screen "St_Parameter" 320x240
   TextField "Text field_13" at 186,102 size 26x12; Text 'Hour'
   TextField "Text field_17" at 122,102 size 34x12; Text 'Second'
   TextField "Text field_10" at 118,88 size 86x16; Text 'Time Shift Setting'
   TextField "Text field_4" at 71,19 size 47x13; Text 'Day (1-31)'
   TextField "Text field_6" at 196,19 size 21x13; Text 'Year'
   TextField "Text field_5" at 119,19 size 61x12; Text 'Month (1-12)'
   TextField "Text field_1" at 6,1 size 143x17; Text 'STATISTIKA PARAMETER'
   TextField "Text field_2" at 9,32 size 62x15; Text 'Date Setting'
   TextField "Text field_3" at 10,65 size 61x15; Text 'Time Setting'
   TextField "Text field_7" at 67,54 size 52x12; Text 'Hour (0-23)'
   TextField "Text field_8" at 119,53 size 59x12; Text 'Minute (0-59)'
   TextField "Text field_9" at 176,53 size 64x12; Text 'Second (0-59)'
   IOField "I/O field_6" at 72,33 size 42x20; FormatPattern 99
      ProcessValue <- "DB_Integer_IDay"
   Button "Button_1" at 256,50 size 57x23; TextOff 'Execute'; TextOn 'OK'
      on Release: ResetBit("Data_Bool1_F_Set Time Day")
      on Press: SetBit("Data_Bool1_F_Set Time Day")
   TextField "Text field_11" at 11,117 size 33x15; Text 'Shift 1'
   TextField "Text field_15" at 49,102 size 26x12; Text 'Hour'
   TextField "Text field_16" at 85,102 size 30x12; Text 'Minute'
   IOField "I/O field_7" at 81,115 size 35x20; FormatPattern 99
      ProcessValue <- "DB_Integer_S1AMinute"
   IOField "I/O field_8" at 119,115 size 35x20; FormatPattern 99
      ProcessValue <- "DB_Integer_S1ASecond"
   TextField "Text field_12" at 160,114 size 17x15; Text 's/d'
   IOField "I/O field_9" at 180,115 size 35x20; FormatPattern 99
      ProcessValue <- "DB_Integer_S1BHour"
   TextField "Text field_14" at 221,102 size 30x12; Text 'Minute'
   TextField "Text field_18" at 256,102 size 34x12; Text 'Second'
   IOField "I/O field_11" at 218,115 size 35x20; FormatPattern 99
      ProcessValue <- "DB_Integer_S1BMinute"
   IOField "I/O field_12" at 256,115 size 35x20; FormatPattern 99
      ProcessValue <- "DB_Integer_S1BSecond"
   TextField "Text field_19" at 10,141 size 33x15; Text 'Shift 2'
   IOField "I/O field_13" at 43,139 size 35x20; FormatPattern 99
      ProcessValue <- "DB_Integer_S2AHour"
   IOField "I/O field_14" at 81,139 size 35x20; FormatPattern 99
      ProcessValue <- "DB_Integer_S2AMinute"
   IOField "I/O field_15" at 119,139 size 35x20; FormatPattern 99
      ProcessValue <- "DB_Integer_S2ASecond"
   TextField "Text field_23" at 160,140 size 17x15; Text 's/d'
   IOField "I/O field_16" at 180,139 size 35x20; FormatPattern 99
      ProcessValue <- "DB_Integer_S2BHour"
   IOField "I/O field_17" at 218,139 size 35x20; FormatPattern 99
      ProcessValue <- "DB_Integer_S2BMinute"
   IOField "I/O field_18" at 256,139 size 35x20; FormatPattern 99
      ProcessValue <- "DB_Integer_S2BSecond"
   TextField "Text field_27" at 9,165 size 33x15; Text 'Shift 3'
   IOField "I/O field_19" at 43,163 size 35x20; FormatPattern 99
      ProcessValue <- "DB_Integer_S3AHour"
   IOField "I/O field_20" at 81,163 size 35x20; FormatPattern 99
      ProcessValue <- "DB_Integer_S3AMinute"
   IOField "I/O field_21" at 119,163 size 35x20; FormatPattern 99
      ProcessValue <- "DB_Integer_S3ASecond"
   TextField "Text field_31" at 160,164 size 17x15; Text 's/d'
   IOField "I/O field_22" at 180,163 size 35x20; FormatPattern 99
      ProcessValue <- "DB_Integer_S3BHour"
   IOField "I/O field_23" at 218,163 size 35x20; FormatPattern 99
      ProcessValue <- "DB_Integer_S3BMinute"
   IOField "I/O field_24" at 256,163 size 35x20; FormatPattern 99
      ProcessValue <- "DB_Integer_S3BSecond"
   IOField "I/O field_10" at 43,115 size 35x20; FormatPattern 99
      ProcessValue <- "DB_Integer_S1AHour"
   IOField "I/O field_1" at 125,33 size 43x20; FormatPattern 99
      ProcessValue <- "DB_Integer_IMonth"
   IOField "I/O field_2" at 180,33 size 52x20; FormatPattern 9999
      ProcessValue <- "DB_Integer_IYear"
   IOField "I/O field_3" at 72,66 size 40x20; FormatPattern 99
      ProcessValue <- "DB_Integer_IHour"
   IOField "I/O field_4" at 129,66 size 40x20; FormatPattern 99
      ProcessValue <- "DB_Integer_IMinute"
   IOField "I/O field_5" at 185,66 size 40x20; FormatPattern 99
      ProcessValue <- "DB_Integer_ISecond"
   IOField "I/O field_25" at 163,1 size 155x23; FormatPattern 9999999999999999999999999999999999999999
      ProcessValue <- "Data_DTL1_Output"
   Button "Button_2" at 138,185 size 57x24; TextOff 'Execute'; TextOn 'OK'
   Button "Button_4" at 3,211 size 35x27; TextOff 'Main Page'; PictureOff "Home"
      on Click: ActivateScreen("Main Page", 0)

screen "Door Open Secret" 320x240
   Button "Button_1" at 100,205 size 120x30; TextOff 'Main Page'
      on Click: ActivateScreen("Main Page", 0)
   Switch "Switch_5" at 100,20 size 107x32; CaptionText 'Switch'; TextOff 'Safety Door On'; TextOn 'Safety Door Off'
      ProcessValue <- "Flag Enable/Disable Error Door Open"
   Switch "Switch_1" at 102,80 size 107x32; TextOff 'Reset'; CaptionText 'Switch'
      ProcessValue <- "AddReject2_DB_CountStop"
   IOField "I/O field_2" at 209,80 size 84x32; FormatPattern 999999999
      ProcessValue <- "AddReject2_DB_Countaddrej"

screen "St_Error Counter" 320x240
   TextField "Text field_13" at 244,51 size 70x129; Text 'Text'
   TextField "Text field_37" at 7,163 size 21x17; Text '8'
   IOField "I/O field_24" at 219,163 size 26x17; FormatPattern 999
      ProcessValue <- "Data_DTLData_DTL_Door Open[0].SECOND"
   IOField "I/O field_25" at 195,163 size 25x17; FormatPattern 999
      ProcessValue <- "Data_DTLData_DTL_Door Open[0].MINUTE"
   IOField "I/O field_26" at 171,163 size 25x17; FormatPattern 999
      ProcessValue <- "Data_DTLData_DTL_Door Open[0].HOUR"
   TextField "Text field_38" at 27,163 size 145x17; Text 'Door Open'
   IOField "I/O field_13" at 219,131 size 26x17; FormatPattern 999
      ProcessValue <- "Data_DTLData_DTL_Press Low[0].SECOND"
   IOField "I/O field_14" at 195,131 size 25x17; FormatPattern 999
      ProcessValue <- "Data_DTLData_DTL_Press Low[0].MINUTE"
   IOField "I/O field_15" at 171,131 size 25x17; FormatPattern 999
      ProcessValue <- "Data_DTLData_DTL_Press Low[0].HOUR"
   TextField "Text field_7" at 27,131 size 145x17; Text 'Pressure Low'
   TextField "Text field_35" at 7,147 size 21x17; Text '7'
   TextField "Text field_34" at 7,131 size 21x17; Text '6'
   TextField "Text field_33" at 7,115 size 21x17; Text '5'
   TextField "Text field_32" at 7,99 size 21x17; Text '4'
   TextField "Text field_31" at 7,83 size 21x17; Text '3'
   TextField "Text field_30" at 7,67 size 21x17; Text '2'
   TextField "Text field_29" at 7,51 size 21x17; Text '1'
   TextField "Text field_28" at 7,35 size 21x17; Text 'No'
   IOField "I/O field_8" at 219,147 size 26x17; FormatPattern 999
      ProcessValue <- "Data_DTLData_DTL_RS Pneu Er.SECOND"
   IOField "I/O field_16" at 195,147 size 25x17; FormatPattern 999
      ProcessValue <- "Data_DTLData_DTL_RS Pneu Er.MINUTE"
   IOField "I/O field_17" at 171,147 size 25x17; FormatPattern 999
      ProcessValue <- "Data_DTLData_DTL_RS Pneu Er.HOUR"
   IOField "I/O field_21" at 219,83 size 26x17; FormatPattern 999
      ProcessValue <- "Data_DTLData_DTL_Imaje Not In Position[0].SECOND"
   IOField "I/O field_22" at 195,83 size 25x17; FormatPattern 999
      ProcessValue <- "Data_DTLData_DTL_Imaje Not In Position[0].MINUTE"
   IOField "I/O field_23" at 171,83 size 25x17; FormatPattern 999
      ProcessValue <- "Data_DTLData_DTL_Imaje Not In Position[0].HOUR"
   TextField "Text field_25" at 27,83 size 145x17; Text 'Imaje Not In Position'
   IOField "I/O field_18" at 219,67 size 26x17; FormatPattern 999
      ProcessValue <- "Data_DTLData_DTL_Paper R Out[0].SECOND"
   IOField "I/O field_19" at 195,67 size 25x17; FormatPattern 999
      ProcessValue <- "Data_DTLData_DTL_Paper R Out[0].MINUTE"
   IOField "I/O field_20" at 171,67 size 25x17; FormatPattern 999
      ProcessValue <- "Data_DTLData_DTL_Paper R Out[0].HOUR"
   TextField "Text field_22" at 27,67 size 145x17; Text 'Imaje Paper Or Ribbon Out'
   TextField "Text field_2" at 171,35 size 25x17; Text 'Hour'
   IOField "I/O field_10" at 219,115 size 26x17; FormatPattern 999
      ProcessValue <- "Data_DTLData_DTL_Sloft Jam1.SECOND"
   IOField "I/O field_11" at 195,115 size 25x17; FormatPattern 999
      ProcessValue <- "Data_DTLData_DTL_Sloft Jam1.MINUTE"
   IOField "I/O field_12" at 171,115 size 25x17; FormatPattern 999
      ProcessValue <- "Data_DTLData_DTL_Sloft Jam1.HOUR"
   IOField "I/O field_4" at 219,99 size 26x17; FormatPattern 999
      ProcessValue <- "Data_DTLData_DTL_Always bad Read[0].SECOND"
   IOField "I/O field_5" at 195,99 size 25x17; FormatPattern 999
      ProcessValue <- "Data_DTLData_DTL_Always bad Read[0].MINUTE"
   IOField "I/O field_9" at 171,99 size 25x17; FormatPattern 999
      ProcessValue <- "Data_DTLData_DTL_Always bad Read[0].HOUR"
   TextField "Text field_12" at 219,35 size 26x17; Text 'Sec'
   TextField "Text field_11" at 195,35 size 25x17; Text 'Min'
   IOField "I/O field_2" at 219,51 size 26x17; FormatPattern 999
      ProcessValue <- "Data_DTLData_DTL_Imaje Er.SECOND"
   IOField "I/O field_1" at 195,51 size 25x17; FormatPattern 999
      ProcessValue <- "Data_DTLData_DTL_Imaje Er.MINUTE"
   TextField "Text field_3" at 27,35 size 145x17; Text 'Error Counter'
   TextField "Text field_4" at 27,51 size 145x17; Text 'System Imaje Error'
   TextField "Text field_5" at 27,99 size 145x17; Text 'Always Bad Read Sloft'
   IOField "I/O field_3" at 171,51 size 25x17; FormatPattern 999
      ProcessValue <- "Data_DTLData_DTL_Imaje Er.HOUR"
   TextField "Text field_9" at 120,17 size 18x13; Text 'S/D'
   TextField "Text field_1" at 3,0 size 197x18; Text 'CURRENT SHIFT (Error Counter)'
   TextField "Text field_36" at 260,0 size 57x15; Text 'Page 3 of 3'
   Button "Button_1" at 46,217 size 90x21; TextOff 'Statistic Data'
      on Click: ActivateScreen("St_Data Statistic", 0)
   Button "Button_3" at 1,218 size 41x20; TextOff 'Main Page'; PictureOff "Home"
      on Click: ActivateScreen("Main Page", 0)
   Button "Button_4" at 151,217 size 80x21; TextOff '<-- Back Page'; TextOn 'Page 2'
      on Click: ActivateScreen("St_Time machine data", 0)
   TextField "Text field_10" at 27,182 size 145x17; Text 'Downstream Jammed'
   IOField "I/O field_30" at 171,182 size 25x17; FormatPattern 999
      ProcessValue <- "Data_DTLData_DTL_Down Stop.HOUR"
   IOField "I/O field_31" at 195,182 size 25x17; FormatPattern 999
      ProcessValue <- "Data_DTLData_DTL_Down Stop.MINUTE"
   IOField "I/O field_32" at 219,182 size 26x17; FormatPattern 999
      ProcessValue <- "Data_DTLData_DTL_Down Stop.SECOND"
   TextField "Text field_14" at 244,182 size 70x17; Text 'Warning'
   IOField "I/O field_6" at 6,17 size 109x15; FormatPattern 9999999999999999999999999999999999999999
      ProcessValue <- "Data_DTL1_Cur_ShiftA"
   IOField "I/O field_7" at 143,17 size 109x15; FormatPattern 9999999999999999999999999999999999999999
      ProcessValue <- "Data_DTL1_Cur_ShiftB"
   TextField "Text field_15" at 263,115 size 7x15; Text ':'
   TextField "Text field_17" at 287,115 size 7x15; Text ':'
   IOField "I/O field_33" at 245,116 size 21x15; FormatPattern 999
      ProcessValue <- "Data_DTLData_DTL_Total Detail Error[0].HOUR"
   IOField "I/O field_34" at 268,116 size 21x15; FormatPattern 999
      ProcessValue <- "Data_DTLData_DTL_Total Detail Error[0].MINUTE"
   IOField "I/O field_35" at 291,116 size 21x15; FormatPattern 999
      ProcessValue <- "Data_DTLData_DTL_Total Detail Error[0].SECOND"
   TextField "Text field_16" at 244,35 size 70x17; Text 'Total (H:M:S)'
   TextField "Text field_8" at 27,115 size 145x17; Text 'Bundle Jammed'
   TextField "Text field_18" at 27,147 size 145x17; Text 'Reed Swicth pneumatic Error'
   IOField "I/O field_27" at 253,16 size 66x17; FormatPattern ????????
      ProcessValue <- "Data_String_sDT_Machine id"

screen "ST_Error Counter_1" 320x240
   TextField "Text field_13" at 244,51 size 70x129; Text 'Text'
   TextField "Text field_37" at 7,163 size 21x17; Text '8'
   IOField "I/O field_24" at 219,163 size 26x17; FormatPattern 999
      ProcessValue <- "Data_DTLData_DTL_Door Open[1].SECOND"
   IOField "I/O field_25" at 195,163 size 25x17; FormatPattern 999
      ProcessValue <- "Data_DTLData_DTL_Door Open[1].MINUTE"
   IOField "I/O field_26" at 171,163 size 25x17; FormatPattern 999
      ProcessValue <- "Data_DTLData_DTL_Door Open[1].HOUR"
   TextField "Text field_38" at 27,163 size 145x17; Text 'Door Open'
   IOField "I/O field_13" at 219,131 size 26x17; FormatPattern 999
      ProcessValue <- "Data_DTLData_DTL_Press Low[1].SECOND"
   IOField "I/O field_14" at 195,131 size 25x17; FormatPattern 999
      ProcessValue <- "Data_DTLData_DTL_Press Low[1].MINUTE"
   IOField "I/O field_15" at 171,131 size 25x17; FormatPattern 999
      ProcessValue <- "Data_DTLData_DTL_Press Low[1].HOUR"
   TextField "Text field_7" at 27,131 size 145x17; Text 'Pressure Low'
   TextField "Text field_35" at 7,147 size 21x17; Text '7'
   TextField "Text field_34" at 7,131 size 21x17; Text '6'
   TextField "Text field_33" at 7,115 size 21x17; Text '5'
   TextField "Text field_32" at 7,99 size 21x17; Text '4'
   TextField "Text field_31" at 7,83 size 21x17; Text '3'
   TextField "Text field_30" at 7,67 size 21x17; Text '2'
   TextField "Text field_29" at 7,51 size 21x17; Text '1'
   TextField "Text field_28" at 7,35 size 21x17; Text 'No'
   IOField "I/O field_8" at 219,147 size 26x17; FormatPattern 999
      ProcessValue <- "Data_DTLData_DTL_RS Pneu Er_1.SECOND"
   IOField "I/O field_16" at 195,147 size 25x17; FormatPattern 999
      ProcessValue <- "Data_DTLData_DTL_RS Pneu Er_1.MINUTE"
   IOField "I/O field_17" at 171,147 size 25x17; FormatPattern 999
      ProcessValue <- "Data_DTLData_DTL_RS Pneu Er_1.HOUR"
   IOField "I/O field_21" at 219,83 size 26x17; FormatPattern 999
      ProcessValue <- "Data_DTLData_DTL_Imaje Not In Position[1].SECOND"
   IOField "I/O field_22" at 195,83 size 25x17; FormatPattern 999
      ProcessValue <- "Data_DTLData_DTL_Imaje Not In Position[1].MINUTE"
   IOField "I/O field_23" at 171,83 size 25x17; FormatPattern 999
      ProcessValue <- "Data_DTLData_DTL_Imaje Not In Position[1].HOUR"
   TextField "Text field_25" at 27,83 size 145x17; Text 'Imaje Not In Position'
   IOField "I/O field_18" at 219,67 size 26x17; FormatPattern 999
      ProcessValue <- "Data_DTLData_DTL_Paper R Out[1].SECOND"
   IOField "I/O field_19" at 195,67 size 25x17; FormatPattern 999
      ProcessValue <- "Data_DTLData_DTL_Paper R Out[1].MINUTE"
   IOField "I/O field_20" at 171,67 size 25x17; FormatPattern 999
      ProcessValue <- "Data_DTLData_DTL_Paper R Out[1].HOUR"
   TextField "Text field_22" at 27,67 size 145x17; Text 'Imaje Paper Or Ribbon Out'
   TextField "Text field_2" at 171,35 size 25x17; Text 'Hour'
   IOField "I/O field_10" at 219,115 size 26x17; FormatPattern 999
      ProcessValue <- "Data_DTLData_DTL_Sloft Jam1_1.SECOND"
   IOField "I/O field_11" at 195,115 size 25x17; FormatPattern 999
      ProcessValue <- "Data_DTLData_DTL_Sloft Jam1_1.MINUTE"
   IOField "I/O field_12" at 171,115 size 25x17; FormatPattern 999
      ProcessValue <- "Data_DTLData_DTL_Sloft Jam1_1.HOUR"
   IOField "I/O field_4" at 219,99 size 26x17; FormatPattern 999
      ProcessValue <- "Data_DTLData_DTL_Always bad Read[1].SECOND"
   IOField "I/O field_5" at 195,99 size 25x17; FormatPattern 999
      ProcessValue <- "Data_DTLData_DTL_Always bad Read[1].MINUTE"
   IOField "I/O field_9" at 171,99 size 25x17; FormatPattern 999
      ProcessValue <- "Data_DTLData_DTL_Always bad Read[1].HOUR"
   TextField "Text field_12" at 219,35 size 26x17; Text 'Sec'
   TextField "Text field_11" at 195,35 size 25x17; Text 'Min'
   IOField "I/O field_2" at 219,51 size 26x17; FormatPattern 999
      ProcessValue <- "Data_DTLData_DTL_Imaje Er_1.SECOND"
   IOField "I/O field_1" at 195,51 size 25x17; FormatPattern 999
      ProcessValue <- "Data_DTLData_DTL_Imaje Er_1.MINUTE"
   TextField "Text field_3" at 27,35 size 145x17; Text 'Error Counter'
   TextField "Text field_4" at 27,51 size 145x17; Text 'System Imaje Error'
   TextField "Text field_5" at 27,99 size 145x17; Text 'Always Bad Read Sloft'
   IOField "I/O field_3" at 171,51 size 25x17; FormatPattern 999
      ProcessValue <- "Data_DTLData_DTL_Imaje Er_1.HOUR"
   TextField "Text field_9" at 120,17 size 18x13; Text 'S/D'
   TextField "Text field_1" at 3,0 size 159x18; Text 'CURRENT SHIFT MINUS 1'
   TextField "Text field_36" at 260,0 size 57x15; Text 'Page 3 of 3'
   Button "Button_1" at 46,217 size 90x21; TextOff 'Statistic Data'
      on Click: ActivateScreen("St_Data Statistic", 0)
   Button "Button_3" at 1,218 size 41x20; TextOff 'Main Page'; PictureOff "Home"
      on Click: ActivateScreen("Main Page", 0)
   Button "Button_4" at 151,217 size 80x21; TextOff '<-- Back Page'; TextOn 'Page 2'
      on Click: ActivateScreen("St_Time machine data_1", 0)
   TextField "Text field_10" at 27,182 size 145x17; Text 'Downstream Jammed'
   IOField "I/O field_30" at 171,182 size 25x17; FormatPattern 999
      ProcessValue <- "Data_DTLData_DTL_Down Stop_1.HOUR"
   IOField "I/O field_31" at 195,182 size 25x17; FormatPattern 999
      ProcessValue <- "Data_DTLData_DTL_Down Stop_1.MINUTE"
   IOField "I/O field_32" at 219,182 size 26x17; FormatPattern 999
      ProcessValue <- "Data_DTLData_DTL_Down Stop_1.SECOND"
   TextField "Text field_14" at 244,182 size 70x17; Text 'Warning'
   IOField "I/O field_7" at 143,17 size 109x15; FormatPattern 9999999999999999999999999999999999999999
      ProcessValue <- "Data_DTL1_Cur_ShiftB_1"
   IOField "I/O field_6" at 6,17 size 109x15; FormatPattern 9999999999999999999999999999999999999999
      ProcessValue <- "Data_DTL1_Cur_ShiftA_1"
   TextField "Text field_15" at 263,115 size 7x15; Text ':'
   TextField "Text field_17" at 287,115 size 7x15; Text ':'
   IOField "I/O field_33" at 245,116 size 21x15; FormatPattern 999
      ProcessValue <- "Data_DTLData_DTL_Total Detail Error[1].HOUR"
   IOField "I/O field_34" at 268,116 size 21x15; FormatPattern 999
      ProcessValue <- "Data_DTLData_DTL_Total Detail Error[1].MINUTE"
   IOField "I/O field_35" at 291,116 size 21x15; FormatPattern 999
      ProcessValue <- "Data_DTLData_DTL_Total Detail Error[1].SECOND"
   TextField "Text field_16" at 244,35 size 70x17; Text 'Total (H:M:S)'
   TextField "Text field_8" at 27,115 size 145x17; Text 'Bundle Jammed'
   TextField "Text field_18" at 27,147 size 145x17; Text 'Reed Swicth pneumatic Error'
   IOField "I/O field_27" at 253,16 size 66x17; FormatPattern ????????
      ProcessValue <- "Data_String_sDT_Machine id"

screen "St_Error Counter_2" 320x240
   TextField "Text field_13" at 244,51 size 70x129; Text 'Text'
   TextField "Text field_37" at 7,163 size 21x17; Text '8'
   IOField "I/O field_24" at 219,163 size 26x17; FormatPattern 999
      ProcessValue <- "Data_DTLData_DTL_Door Open[2].SECOND"
   IOField "I/O field_25" at 195,163 size 25x17; FormatPattern 999
      ProcessValue <- "Data_DTLData_DTL_Door Open[2].MINUTE"
   IOField "I/O field_26" at 171,163 size 25x17; FormatPattern 999
      ProcessValue <- "Data_DTLData_DTL_Door Open[2].HOUR"
   TextField "Text field_38" at 27,163 size 145x17; Text 'Door Open'
   IOField "I/O field_13" at 219,131 size 26x17; FormatPattern 999
      ProcessValue <- "Data_DTLData_DTL_Press Low[2].SECOND"
   IOField "I/O field_14" at 195,131 size 25x17; FormatPattern 999
      ProcessValue <- "Data_DTLData_DTL_Press Low[2].MINUTE"
   IOField "I/O field_15" at 171,131 size 25x17; FormatPattern 999
      ProcessValue <- "Data_DTLData_DTL_Press Low[2].HOUR"
   TextField "Text field_7" at 27,131 size 145x17; Text 'Pressure Low'
   TextField "Text field_35" at 7,147 size 21x17; Text '7'
   TextField "Text field_34" at 7,131 size 21x17; Text '6'
   TextField "Text field_33" at 7,115 size 21x17; Text '5'
   TextField "Text field_32" at 7,99 size 21x17; Text '4'
   TextField "Text field_31" at 7,83 size 21x17; Text '3'
   TextField "Text field_30" at 7,67 size 21x17; Text '2'
   TextField "Text field_29" at 7,51 size 21x17; Text '1'
   TextField "Text field_28" at 7,35 size 21x17; Text 'No'
   IOField "I/O field_8" at 219,147 size 26x17; FormatPattern 999
      ProcessValue <- "Data_DTLData_DTL_RS Pneu Er_2.SECOND"
   IOField "I/O field_16" at 195,147 size 25x17; FormatPattern 999
      ProcessValue <- "Data_DTLData_DTL_RS Pneu Er_2.MINUTE"
   IOField "I/O field_17" at 171,147 size 25x17; FormatPattern 999
      ProcessValue <- "Data_DTLData_DTL_RS Pneu Er_2.HOUR"
   IOField "I/O field_21" at 219,83 size 26x17; FormatPattern 999
      ProcessValue <- "Data_DTLData_DTL_Imaje Not In Position[2].SECOND"
   IOField "I/O field_22" at 195,83 size 25x17; FormatPattern 999
      ProcessValue <- "Data_DTLData_DTL_Imaje Not In Position[2].MINUTE"
   IOField "I/O field_23" at 171,83 size 25x17; FormatPattern 999
      ProcessValue <- "Data_DTLData_DTL_Imaje Not In Position[2].HOUR"
   TextField "Text field_25" at 27,83 size 145x17; Text 'Imaje Not In Position'
   IOField "I/O field_18" at 219,67 size 26x17; FormatPattern 999
      ProcessValue <- "Data_DTLData_DTL_Paper R Out[2].SECOND"
   IOField "I/O field_19" at 195,67 size 25x17; FormatPattern 999
      ProcessValue <- "Data_DTLData_DTL_Paper R Out[2].MINUTE"
   IOField "I/O field_20" at 171,67 size 25x17; FormatPattern 999
      ProcessValue <- "Data_DTLData_DTL_Paper R Out[2].HOUR"
   TextField "Text field_22" at 27,67 size 145x17; Text 'Imaje Paper Or Ribbon Out'
   TextField "Text field_2" at 171,35 size 25x17; Text 'Hour'
   IOField "I/O field_10" at 219,115 size 26x17; FormatPattern 999
      ProcessValue <- "Data_DTLData_DTL_Sloft Jam1_2.SECOND"
   IOField "I/O field_11" at 195,115 size 25x17; FormatPattern 999
      ProcessValue <- "Data_DTLData_DTL_Sloft Jam1_2.MINUTE"
   IOField "I/O field_12" at 171,115 size 25x17; FormatPattern 999
      ProcessValue <- "Data_DTLData_DTL_Sloft Jam1_2.HOUR"
   IOField "I/O field_4" at 219,99 size 26x17; FormatPattern 999
      ProcessValue <- "Data_DTLData_DTL_Always bad Read[2].SECOND"
   IOField "I/O field_5" at 195,99 size 25x17; FormatPattern 999
      ProcessValue <- "Data_DTLData_DTL_Always bad Read[2].MINUTE"
   IOField "I/O field_9" at 171,99 size 25x17; FormatPattern 999
      ProcessValue <- "Data_DTLData_DTL_Always bad Read[2].HOUR"
   TextField "Text field_12" at 219,35 size 26x17; Text 'Sec'
   TextField "Text field_11" at 195,35 size 25x17; Text 'Min'
   IOField "I/O field_2" at 219,51 size 26x17; FormatPattern 999
      ProcessValue <- "Data_DTLData_DTL_Imaje Er_2.SECOND"
   IOField "I/O field_1" at 195,51 size 25x17; FormatPattern 999
      ProcessValue <- "Data_DTLData_DTL_Imaje Er_2.MINUTE"
   TextField "Text field_3" at 27,35 size 145x17; Text 'Error Counter'
   TextField "Text field_4" at 27,51 size 145x17; Text 'System Imaje Error'
   TextField "Text field_5" at 27,99 size 145x17; Text 'Always Bad Read Sloft'
   IOField "I/O field_3" at 171,51 size 25x17; FormatPattern 999
      ProcessValue <- "Data_DTLData_DTL_Imaje Er_2.HOUR"
   IOField "I/O field_6" at 6,17 size 109x15; FormatPattern 9999999999999999999999999999999999999999
      ProcessValue <- "Data_DTL1_Cur_ShiftA_2"
   TextField "Text field_9" at 120,17 size 18x13; Text 'S/D'
   IOField "I/O field_7" at 143,17 size 109x15; FormatPattern 9999999999999999999999999999999999999999
      ProcessValue <- "Data_DTL1_Cur_ShiftB_2"
   TextField "Text field_1" at 3,0 size 159x18; Text 'CURRENT SHIFT MINUS 2'
   TextField "Text field_36" at 260,0 size 57x15; Text 'Page 3 of 3'
   Button "Button_1" at 46,217 size 90x21; TextOff 'Statistic Data'
      on Click: ActivateScreen("St_Data Statistic", 0)
   Button "Button_3" at 1,218 size 41x20; TextOff 'Main Page'; PictureOff "Home"
      on Click: ActivateScreen("Main Page", 0)
   Button "Button_4" at 151,217 size 80x21; TextOff '<-- Back Page'; TextOn 'Page 2'
      on Click: ActivateScreen("St_Time machine data_2", 0)
   TextField "Text field_10" at 27,182 size 145x17; Text 'Downstream Jammed'
   IOField "I/O field_30" at 171,182 size 25x17; FormatPattern 999
      ProcessValue <- "Data_DTLData_DTL_Down Stop_2.HOUR"
   IOField "I/O field_31" at 195,182 size 25x17; FormatPattern 999
      ProcessValue <- "Data_DTLData_DTL_Down Stop_2.MINUTE"
   IOField "I/O field_32" at 219,182 size 26x17; FormatPattern 999
      ProcessValue <- "Data_DTLData_DTL_Down Stop_2.SECOND"
   TextField "Text field_14" at 244,182 size 70x17; Text 'Warning'
   TextField "Text field_15" at 263,115 size 7x15; Text ':'
   TextField "Text field_17" at 287,115 size 7x15; Text ':'
   IOField "I/O field_33" at 245,116 size 21x15; FormatPattern 999
      ProcessValue <- "Data_DTLData_DTL_Total Detail Error[2].HOUR"
   IOField "I/O field_34" at 268,116 size 21x15; FormatPattern 999
      ProcessValue <- "Data_DTLData_DTL_Total Detail Error[2].MINUTE"
   IOField "I/O field_35" at 291,116 size 21x15; FormatPattern 999
      ProcessValue <- "Data_DTLData_DTL_Total Detail Error[2].SECOND"
   TextField "Text field_16" at 244,35 size 70x17; Text 'Total (H:M:S)'
   TextField "Text field_8" at 27,115 size 145x17; Text 'Bundle Jammed'
   TextField "Text field_18" at 27,147 size 145x17; Text 'Reed Swicth pneumatic Error'
   IOField "I/O field_27" at 253,16 size 66x17; FormatPattern ????????
      ProcessValue <- "Data_String_sDT_Machine id"

screen "St_Error Counter_3" 320x240
   TextField "Text field_13" at 244,51 size 70x129; Text 'Text'
   TextField "Text field_37" at 7,163 size 21x17; Text '8'
   IOField "I/O field_24" at 219,163 size 26x17; FormatPattern 999
      ProcessValue <- "Data_DTLData_DTL_Door Open[3].SECOND"
   IOField "I/O field_25" at 195,163 size 25x17; FormatPattern 999
      ProcessValue <- "Data_DTLData_DTL_Door Open[3].MINUTE"
   IOField "I/O field_26" at 171,163 size 25x17; FormatPattern 999
      ProcessValue <- "Data_DTLData_DTL_Door Open[3].HOUR"
   TextField "Text field_38" at 27,163 size 145x17; Text 'Door Open'
   IOField "I/O field_13" at 219,131 size 26x17; FormatPattern 999
      ProcessValue <- "Data_DTLData_DTL_Press Low[3].SECOND"
   IOField "I/O field_14" at 195,131 size 25x17; FormatPattern 999
      ProcessValue <- "Data_DTLData_DTL_Press Low[3].MINUTE"
   IOField "I/O field_15" at 171,131 size 25x17; FormatPattern 999
      ProcessValue <- "Data_DTLData_DTL_Press Low[3].HOUR"
   TextField "Text field_7" at 27,131 size 145x17; Text 'Pressure Low'
   TextField "Text field_35" at 7,147 size 21x17; Text '7'
   TextField "Text field_34" at 7,131 size 21x17; Text '6'
   TextField "Text field_33" at 7,115 size 21x17; Text '5'
   TextField "Text field_32" at 7,99 size 21x17; Text '4'
   TextField "Text field_31" at 7,83 size 21x17; Text '3'
   TextField "Text field_30" at 7,67 size 21x17; Text '2'
   TextField "Text field_29" at 7,51 size 21x17; Text '1'
   TextField "Text field_28" at 7,35 size 21x17; Text 'No'
   IOField "I/O field_8" at 219,147 size 26x17; FormatPattern 999
      ProcessValue <- "Data_DTLData_DTL_RS Pneu Er_3.SECOND"
   IOField "I/O field_16" at 195,147 size 25x17; FormatPattern 999
      ProcessValue <- "Data_DTLData_DTL_RS Pneu Er_3.MINUTE"
   IOField "I/O field_17" at 171,147 size 25x17; FormatPattern 999
      ProcessValue <- "Data_DTLData_DTL_RS Pneu Er_3.HOUR"
   IOField "I/O field_21" at 219,83 size 26x17; FormatPattern 999
      ProcessValue <- "Data_DTLData_DTL_Imaje Not In Position[3].SECOND"
   IOField "I/O field_22" at 195,83 size 25x17; FormatPattern 999
      ProcessValue <- "Data_DTLData_DTL_Imaje Not In Position[3].MINUTE"
   IOField "I/O field_23" at 171,83 size 25x17; FormatPattern 999
      ProcessValue <- "Data_DTLData_DTL_Imaje Not In Position[3].HOUR"
   TextField "Text field_25" at 27,83 size 145x17; Text 'Imaje Not In Position'
   IOField "I/O field_18" at 219,67 size 26x17; FormatPattern 999
      ProcessValue <- "Data_DTLData_DTL_Paper R Out[3].SECOND"
   IOField "I/O field_19" at 195,67 size 25x17; FormatPattern 999
      ProcessValue <- "Data_DTLData_DTL_Paper R Out[3].MINUTE"
   IOField "I/O field_20" at 171,67 size 25x17; FormatPattern 999
      ProcessValue <- "Data_DTLData_DTL_Paper R Out[3].HOUR"
   TextField "Text field_22" at 27,67 size 145x17; Text 'Imaje Paper Or Ribbon Out'
   TextField "Text field_2" at 171,35 size 25x17; Text 'Hour'
   IOField "I/O field_10" at 219,115 size 26x17; FormatPattern 999
      ProcessValue <- "Data_DTLData_DTL_Sloft Jam1_3.SECOND"
   IOField "I/O field_11" at 195,115 size 25x17; FormatPattern 999
      ProcessValue <- "Data_DTLData_DTL_Sloft Jam1_3.MINUTE"
   IOField "I/O field_12" at 171,115 size 25x17; FormatPattern 999
      ProcessValue <- "Data_DTLData_DTL_Sloft Jam1_3.HOUR"
   IOField "I/O field_4" at 219,99 size 26x17; FormatPattern 999
      ProcessValue <- "Data_DTLData_DTL_Always bad Read[3].SECOND"
   IOField "I/O field_5" at 195,99 size 25x17; FormatPattern 999
      ProcessValue <- "Data_DTLData_DTL_Always bad Read[3].MINUTE"
   IOField "I/O field_9" at 171,99 size 25x17; FormatPattern 999
      ProcessValue <- "Data_DTLData_DTL_Always bad Read[3].HOUR"
   TextField "Text field_12" at 219,35 size 26x17; Text 'Sec'
   TextField "Text field_11" at 195,35 size 25x17; Text 'Min'
   IOField "I/O field_2" at 219,51 size 26x17; FormatPattern 999
      ProcessValue <- "Data_DTLData_DTL_Imaje Er_3.SECOND"
   IOField "I/O field_1" at 195,51 size 25x17; FormatPattern 999
      ProcessValue <- "Data_DTLData_DTL_Imaje Er_3.MINUTE"
   TextField "Text field_3" at 27,35 size 145x17; Text 'Error Counter'
   TextField "Text field_4" at 27,51 size 145x17; Text 'System Imaje Error'
   TextField "Text field_5" at 27,99 size 145x17; Text 'Always Bad Read Sloft'
   IOField "I/O field_3" at 171,51 size 25x17; FormatPattern 999
      ProcessValue <- "Data_DTLData_DTL_Imaje Er_3.HOUR"
   IOField "I/O field_6" at 6,17 size 109x15; FormatPattern 9999999999999999999999999999999999999999
      ProcessValue <- "Data_DTL1_Cur_ShiftA_3"
   TextField "Text field_9" at 120,17 size 18x13; Text 'S/D'
   IOField "I/O field_7" at 143,17 size 109x15; FormatPattern 9999999999999999999999999999999999999999
      ProcessValue <- "Data_DTL1_Cur_ShiftB_3"
   TextField "Text field_1" at 3,0 size 159x18; Text 'CURRENT SHIFT MINUS 3'
   TextField "Text field_36" at 260,0 size 57x15; Text 'Page 3 of 3'
   Button "Button_1" at 46,217 size 90x21; TextOff 'Statistic Data'
      on Click: ActivateScreen("St_Data Statistic", 0)
   Button "Button_3" at 1,218 size 41x20; TextOff 'Main Page'; PictureOff "Home"
      on Click: ActivateScreen("Main Page", 0)
   Button "Button_4" at 151,217 size 80x21; TextOff '<-- Back Page'; TextOn 'Page 2'
      on Click: ActivateScreen("St_Time machine data_3", 0)
   TextField "Text field_10" at 27,182 size 145x17; Text 'Downstream Jammed'
   IOField "I/O field_30" at 171,182 size 25x17; FormatPattern 999
      ProcessValue <- "Data_DTLData_DTL_Down Stop_3.HOUR"
   IOField "I/O field_31" at 195,182 size 25x17; FormatPattern 999
      ProcessValue <- "Data_DTLData_DTL_Down Stop_3.MINUTE"
   IOField "I/O field_32" at 219,182 size 26x17; FormatPattern 999
      ProcessValue <- "Data_DTLData_DTL_Down Stop_3.SECOND"
   TextField "Text field_14" at 244,182 size 70x17; Text 'Warning'
   TextField "Text field_15" at 263,115 size 7x15; Text ':'
   TextField "Text field_17" at 287,115 size 7x15; Text ':'
   IOField "I/O field_33" at 245,116 size 21x15; FormatPattern 999
      ProcessValue <- "Data_DTLData_DTL_Total Detail Error[3].HOUR"
   IOField "I/O field_34" at 268,116 size 21x15; FormatPattern 999
      ProcessValue <- "Data_DTLData_DTL_Total Detail Error[3].MINUTE"
   IOField "I/O field_35" at 291,116 size 21x15; FormatPattern 999
      ProcessValue <- "Data_DTLData_DTL_Total Detail Error[3].SECOND"
   TextField "Text field_16" at 244,35 size 70x17; Text 'Total (H:M:S)'
   TextField "Text field_8" at 27,115 size 145x17; Text 'Bundle Jammed'
   TextField "Text field_18" at 27,147 size 145x17; Text 'Reed Swicth pneumatic Error'
   IOField "I/O field_27" at 253,16 size 66x17; FormatPattern ????????
      ProcessValue <- "Data_String_sDT_Machine id"

screen "St_Error Counter_4" 320x240
   TextField "Text field_13" at 244,51 size 70x129; Text 'Text'
   TextField "Text field_37" at 7,163 size 21x17; Text '8'
   IOField "I/O field_24" at 219,163 size 26x17; FormatPattern 999
      ProcessValue <- "Data_DTLData_DTL_Door Open[4].SECOND"
   IOField "I/O field_25" at 195,163 size 25x17; FormatPattern 999
      ProcessValue <- "Data_DTLData_DTL_Door Open[4].MINUTE"
   IOField "I/O field_26" at 171,163 size 25x17; FormatPattern 999
      ProcessValue <- "Data_DTLData_DTL_Door Open[4].HOUR"
   TextField "Text field_38" at 27,163 size 145x17; Text 'Door Open'
   IOField "I/O field_13" at 219,131 size 26x17; FormatPattern 999
      ProcessValue <- "Data_DTLData_DTL_Press Low[4].SECOND"
   IOField "I/O field_14" at 195,131 size 25x17; FormatPattern 999
      ProcessValue <- "Data_DTLData_DTL_Press Low[4].MINUTE"
   IOField "I/O field_15" at 171,131 size 25x17; FormatPattern 999
      ProcessValue <- "Data_DTLData_DTL_Press Low[4].HOUR"
   TextField "Text field_7" at 27,131 size 145x17; Text 'Pressure Low'
   TextField "Text field_35" at 7,147 size 21x17; Text '7'
   TextField "Text field_34" at 7,131 size 21x17; Text '6'
   TextField "Text field_33" at 7,115 size 21x17; Text '5'
   TextField "Text field_32" at 7,99 size 21x17; Text '4'
   TextField "Text field_31" at 7,83 size 21x17; Text '3'
   TextField "Text field_30" at 7,67 size 21x17; Text '2'
   TextField "Text field_29" at 7,51 size 21x17; Text '1'
   TextField "Text field_28" at 7,35 size 21x17; Text 'No'
   IOField "I/O field_8" at 219,147 size 26x17; FormatPattern 999
      ProcessValue <- "Data_DTLData_DTL_RS Pneu Er_4.SECOND"
   IOField "I/O field_16" at 195,147 size 25x17; FormatPattern 999
      ProcessValue <- "Data_DTLData_DTL_RS Pneu Er_4.MINUTE"
   IOField "I/O field_17" at 171,147 size 25x17; FormatPattern 999
      ProcessValue <- "Data_DTLData_DTL_RS Pneu Er_4.HOUR"
   IOField "I/O field_21" at 219,83 size 26x17; FormatPattern 999
      ProcessValue <- "Data_DTLData_DTL_Imaje Not In Position[4].SECOND"
   IOField "I/O field_22" at 195,83 size 25x17; FormatPattern 999
      ProcessValue <- "Data_DTLData_DTL_Imaje Not In Position[4].MINUTE"
   IOField "I/O field_23" at 171,83 size 25x17; FormatPattern 999
      ProcessValue <- "Data_DTLData_DTL_Imaje Not In Position[4].HOUR"
   TextField "Text field_25" at 27,83 size 145x17; Text 'Imaje Not In Position'
   IOField "I/O field_18" at 219,67 size 26x17; FormatPattern 999
      ProcessValue <- "Data_DTLData_DTL_Paper R Out[4].SECOND"
   IOField "I/O field_19" at 195,67 size 25x17; FormatPattern 999
      ProcessValue <- "Data_DTLData_DTL_Paper R Out[4].MINUTE"
   IOField "I/O field_20" at 171,67 size 25x17; FormatPattern 999
      ProcessValue <- "Data_DTLData_DTL_Paper R Out[4].HOUR"
   TextField "Text field_22" at 27,67 size 145x17; Text 'Imaje Paper Or Ribbon Out'
   TextField "Text field_2" at 171,35 size 25x17; Text 'Hour'
   IOField "I/O field_10" at 219,115 size 26x17; FormatPattern 999
      ProcessValue <- "Data_DTLData_DTL_Sloft Jam1_4.SECOND"
   IOField "I/O field_11" at 195,115 size 25x17; FormatPattern 999
      ProcessValue <- "Data_DTLData_DTL_Sloft Jam1_4.MINUTE"
   IOField "I/O field_12" at 171,115 size 25x17; FormatPattern 999
      ProcessValue <- "Data_DTLData_DTL_Sloft Jam1_4.HOUR"
   IOField "I/O field_4" at 219,99 size 26x17; FormatPattern 999
      ProcessValue <- "Data_DTLData_DTL_Always bad Read[4].SECOND"
   IOField "I/O field_5" at 195,99 size 25x17; FormatPattern 999
      ProcessValue <- "Data_DTLData_DTL_Always bad Read[4].MINUTE"
   IOField "I/O field_9" at 171,99 size 25x17; FormatPattern 999
      ProcessValue <- "Data_DTLData_DTL_Always bad Read[4].HOUR"
   TextField "Text field_12" at 219,35 size 26x17; Text 'Sec'
   TextField "Text field_11" at 195,35 size 25x17; Text 'Min'
   IOField "I/O field_2" at 219,51 size 26x17; FormatPattern 999
      ProcessValue <- "Data_DTLData_DTL_Imaje Er_4.SECOND"
   IOField "I/O field_1" at 195,51 size 25x17; FormatPattern 999
      ProcessValue <- "Data_DTLData_DTL_Imaje Er_4.MINUTE"
   TextField "Text field_3" at 27,35 size 145x17; Text 'Error Counter'
   TextField "Text field_4" at 27,51 size 145x17; Text 'System Imaje Error'
   TextField "Text field_5" at 27,99 size 145x17; Text 'Always Bad Read Sloft'
   IOField "I/O field_3" at 171,51 size 25x17; FormatPattern 999
      ProcessValue <- "Data_DTLData_DTL_Imaje Er_4.HOUR"
   IOField "I/O field_6" at 6,17 size 109x15; FormatPattern 9999999999999999999999999999999999999999
      ProcessValue <- "Data_DTL1_Cur_ShiftA_4"
   TextField "Text field_9" at 120,17 size 18x13; Text 'S/D'
   IOField "I/O field_7" at 143,17 size 109x15; FormatPattern 9999999999999999999999999999999999999999
      ProcessValue <- "Data_DTL1_Cur_ShiftB_4"
   TextField "Text field_1" at 3,0 size 155x18; Text 'CURRENT SHIFT MINUS 4'
   TextField "Text field_36" at 260,0 size 57x15; Text 'Page 3 of 3'
   Button "Button_1" at 46,217 size 90x21; TextOff 'Statistic Data'
      on Click: ActivateScreen("St_Data Statistic", 0)
   Button "Button_3" at 1,218 size 41x20; TextOff 'Main Page'; PictureOff "Home"
      on Click: ActivateScreen("Main Page", 0)
   Button "Button_4" at 151,217 size 80x21; TextOff '<-- Back Page'; TextOn 'Page 2'
      on Click: ActivateScreen("St_Time machine data_4", 0)
   TextField "Text field_10" at 27,183 size 145x17; Text 'Downstream Jammed'
   IOField "I/O field_30" at 171,183 size 25x17; FormatPattern 999
      ProcessValue <- "Data_DTLData_DTL_Down Stop_4.HOUR"
   IOField "I/O field_31" at 195,183 size 25x17; FormatPattern 999
      ProcessValue <- "Data_DTLData_DTL_Down Stop_4.MINUTE"
   IOField "I/O field_32" at 219,183 size 26x17; FormatPattern 999
      ProcessValue <- "Data_DTLData_DTL_Down Stop_4.SECOND"
   TextField "Text field_14" at 244,183 size 70x17; Text 'Warning'
   TextField "Text field_15" at 263,115 size 7x15; Text ':'
   TextField "Text field_17" at 287,115 size 7x15; Text ':'
   IOField "I/O field_33" at 245,116 size 21x15; FormatPattern 999
      ProcessValue <- "Data_DTLData_DTL_Total Detail Error[4].HOUR"
   IOField "I/O field_34" at 268,116 size 21x15; FormatPattern 999
      ProcessValue <- "Data_DTLData_DTL_Total Detail Error[4].MINUTE"
   IOField "I/O field_35" at 291,116 size 21x15; FormatPattern 999
      ProcessValue <- "Data_DTLData_DTL_Total Detail Error[4].SECOND"
   TextField "Text field_16" at 244,35 size 70x17; Text 'Total (H:M:S)'
   TextField "Text field_8" at 27,115 size 145x17; Text 'Bundle Jammed'
   TextField "Text field_18" at 27,147 size 145x17; Text 'Reed Swicth pneumatic Error'
   IOField "I/O field_27" at 253,16 size 66x17; FormatPattern ????????
      ProcessValue <- "Data_String_sDT_Machine id"

screen "St_Error Counter_5" 320x240
   TextField "Text field_13" at 244,51 size 70x129; Text 'Text'
   TextField "Text field_37" at 7,163 size 21x17; Text '8'
   IOField "I/O field_24" at 219,163 size 26x17; FormatPattern 999
      ProcessValue <- "Data_DTLData_DTL_Door Open[5].SECOND"
   IOField "I/O field_25" at 195,163 size 25x17; FormatPattern 999
      ProcessValue <- "Data_DTLData_DTL_Door Open[5].MINUTE"
   IOField "I/O field_26" at 171,163 size 25x17; FormatPattern 999
      ProcessValue <- "Data_DTLData_DTL_Door Open[5].HOUR"
   TextField "Text field_38" at 27,163 size 145x17; Text 'Door Open'
   IOField "I/O field_13" at 219,131 size 26x17; FormatPattern 999
      ProcessValue <- "Data_DTLData_DTL_Press Low[5].SECOND"
   IOField "I/O field_14" at 195,131 size 25x17; FormatPattern 999
      ProcessValue <- "Data_DTLData_DTL_Press Low[5].MINUTE"
   IOField "I/O field_15" at 171,131 size 25x17; FormatPattern 999
      ProcessValue <- "Data_DTLData_DTL_Press Low[5].HOUR"
   TextField "Text field_7" at 27,131 size 145x17; Text 'Pressure Low'
   TextField "Text field_35" at 7,147 size 21x17; Text '7'
   TextField "Text field_34" at 7,131 size 21x17; Text '6'
   TextField "Text field_33" at 7,115 size 21x17; Text '5'
   TextField "Text field_32" at 7,99 size 21x17; Text '4'
   TextField "Text field_31" at 7,83 size 21x17; Text '3'
   TextField "Text field_30" at 7,67 size 21x17; Text '2'
   TextField "Text field_29" at 7,51 size 21x17; Text '1'
   TextField "Text field_28" at 7,35 size 21x17; Text 'No'
   IOField "I/O field_8" at 219,147 size 26x17; FormatPattern 999
      ProcessValue <- "Data_DTLData_DTL_RS Pneu Er_5.SECOND"
   IOField "I/O field_16" at 195,147 size 25x17; FormatPattern 999
      ProcessValue <- "Data_DTLData_DTL_RS Pneu Er_5.MINUTE"
   IOField "I/O field_17" at 171,147 size 25x17; FormatPattern 999
      ProcessValue <- "Data_DTLData_DTL_RS Pneu Er_5.HOUR"
   IOField "I/O field_21" at 219,83 size 26x17; FormatPattern 999
      ProcessValue <- "Data_DTLData_DTL_Imaje Not In Position[5].SECOND"
   IOField "I/O field_22" at 195,83 size 25x17; FormatPattern 999
      ProcessValue <- "Data_DTLData_DTL_Imaje Not In Position[5].MINUTE"
   IOField "I/O field_23" at 171,83 size 25x17; FormatPattern 999
      ProcessValue <- "Data_DTLData_DTL_Imaje Not In Position[5].HOUR"
   TextField "Text field_25" at 27,83 size 145x17; Text 'Imaje Not In Position'
   IOField "I/O field_18" at 219,67 size 26x17; FormatPattern 999
      ProcessValue <- "Data_DTLData_DTL_Paper R Out[5].SECOND"
   IOField "I/O field_19" at 195,67 size 25x17; FormatPattern 999
      ProcessValue <- "Data_DTLData_DTL_Paper R Out[5].MINUTE"
   IOField "I/O field_20" at 171,67 size 25x17; FormatPattern 999
      ProcessValue <- "Data_DTLData_DTL_Paper R Out[5].HOUR"
   TextField "Text field_22" at 27,67 size 145x17; Text 'Imaje Paper Or Ribbon Out'
   TextField "Text field_2" at 171,35 size 25x17; Text 'Hour'
   IOField "I/O field_10" at 219,115 size 26x17; FormatPattern 999
      ProcessValue <- "Data_DTLData_DTL_Sloft Jam1_5.SECOND"
   IOField "I/O field_11" at 195,115 size 25x17; FormatPattern 999
      ProcessValue <- "Data_DTLData_DTL_Sloft Jam1_5.MINUTE"
   IOField "I/O field_12" at 171,115 size 25x17; FormatPattern 999
      ProcessValue <- "Data_DTLData_DTL_Sloft Jam1_5.HOUR"
   IOField "I/O field_4" at 219,99 size 26x17; FormatPattern 999
      ProcessValue <- "Data_DTLData_DTL_Always bad Read[5].SECOND"
   IOField "I/O field_5" at 195,99 size 25x17; FormatPattern 999
      ProcessValue <- "Data_DTLData_DTL_Always bad Read[5].MINUTE"
   IOField "I/O field_9" at 171,99 size 25x17; FormatPattern 999
      ProcessValue <- "Data_DTLData_DTL_Always bad Read[5].HOUR"
   TextField "Text field_12" at 219,35 size 26x17; Text 'Sec'
   TextField "Text field_11" at 195,35 size 25x17; Text 'Min'
   IOField "I/O field_2" at 219,51 size 26x17; FormatPattern 999
      ProcessValue <- "Data_DTLData_DTL_Imaje Er_5.SECOND"
   IOField "I/O field_1" at 195,51 size 25x17; FormatPattern 999
      ProcessValue <- "Data_DTLData_DTL_Imaje Er_5.MINUTE"
   TextField "Text field_3" at 27,35 size 145x17; Text 'Error Counter'
   TextField "Text field_4" at 27,51 size 145x17; Text 'System Imaje Error'
   TextField "Text field_5" at 27,99 size 145x17; Text 'Always Bad Read Sloft'
   IOField "I/O field_3" at 171,51 size 25x17; FormatPattern 999
      ProcessValue <- "Data_DTLData_DTL_Imaje Er_5.HOUR"
   IOField "I/O field_6" at 6,17 size 109x15; FormatPattern 9999999999999999999999999999999999999999
      ProcessValue <- "Data_DTL1_Cur_ShiftA_5"
   TextField "Text field_9" at 120,17 size 18x13; Text 'S/D'
   IOField "I/O field_7" at 143,17 size 109x15; FormatPattern 9999999999999999999999999999999999999999
      ProcessValue <- "Data_DTL1_Cur_ShiftB_5"
   TextField "Text field_1" at 3,0 size 155x18; Text 'CURRENT SHIFT MINUS 5'
   TextField "Text field_36" at 260,0 size 57x15; Text 'Page 3 of 3'
   Button "Button_1" at 46,217 size 90x21; TextOff 'Statistic Data'
      on Click: ActivateScreen("St_Data Statistic", 0)
   Button "Button_3" at 1,218 size 41x20; TextOff 'Main Page'; PictureOff "Home"
      on Click: ActivateScreen("Main Page", 0)
   Button "Button_4" at 151,217 size 80x21; TextOff '<-- Back Page'; TextOn 'Page 2'
      on Click: ActivateScreen("St_Time machine data_5", 0)
   TextField "Text field_10" at 27,182 size 145x17; Text 'Downstream Jammed'
   IOField "I/O field_30" at 171,182 size 25x17; FormatPattern 999
      ProcessValue <- "Data_DTLData_DTL_Down Stop_5.HOUR"
   IOField "I/O field_31" at 195,182 size 25x17; FormatPattern 999
      ProcessValue <- "Data_DTLData_DTL_Down Stop_5.MINUTE"
   IOField "I/O field_32" at 219,182 size 26x17; FormatPattern 999
      ProcessValue <- "Data_DTLData_DTL_Down Stop_5.SECOND"
   TextField "Text field_14" at 244,182 size 70x17; Text 'Warning'
   TextField "Text field_16" at 244,35 size 70x17; Text 'Total (H:M:S)'
   TextField "Text field_15" at 263,115 size 7x15; Text ':'
   TextField "Text field_17" at 287,115 size 7x15; Text ':'
   IOField "I/O field_33" at 245,116 size 21x15; FormatPattern 999
      ProcessValue <- "Data_DTLData_DTL_Total Detail Error[5].HOUR"
   IOField "I/O field_34" at 268,116 size 21x15; FormatPattern 999
      ProcessValue <- "Data_DTLData_DTL_Total Detail Error[5].MINUTE"
   IOField "I/O field_35" at 291,116 size 21x15; FormatPattern 999
      ProcessValue <- "Data_DTLData_DTL_Total Detail Error[5].SECOND"
   TextField "Text field_8" at 27,115 size 145x17; Text 'Bundle Jammed'
   TextField "Text field_18" at 27,147 size 145x17; Text 'Reed Swicth pneumatic Error'
   IOField "I/O field_27" at 253,16 size 66x17; FormatPattern ????????
      ProcessValue <- "Data_String_sDT_Machine id"

screen "St_Output Bundled" 320x240
   IOField "I/O field_9" at 228,67 size 87x20; FormatPattern 999.99
      ProcessValue <- "Data_Real_% label Sloft[0]"
   IOField "I/O field_10" at 228,86 size 87x20; FormatPattern 999.99
      ProcessValue <- "Data_Real_% Unlabel Sloft[0]"
   TextField "Text field_1" at 4,0 size 212x18; Text 'CURRENT SHIFT ( Output Bundle )'
   IOField "I/O field_2" at 145,86 size 84x20; FormatPattern 9999999
      ProcessValue <- "Data_IntData_Un label Sloft[0]"
   IOField "I/O field_3" at 145,67 size 84x20; FormatPattern 9999999
      ProcessValue <- "Data_IntData_Label Sloft[0]"
   Button "Button_1" at 101,214 size 128x25; TextOff 'Back To Quantity Data'; TextOn 'Page 1'
      on Click: ActivateScreen("St_Quantity Data", 0)
   IOField "I/O field_6" at 6,17 size 109x15; FormatPattern 9999999999999999999999999999999999999999
      ProcessValue <- "Data_DTL1_Cur_ShiftA"
   TextField "Text field_9" at 120,17 size 18x13; Text 'S/D'
   IOField "I/O field_7" at 143,17 size 109x15; FormatPattern 9999999999999999999999999999999999999999
      ProcessValue <- "Data_DTL1_Cur_ShiftB"
   TextField "Text field_5" at 7,86 size 139x20; Text 'Unlabeled Bundle'
   TextField "Text field_4" at 7,67 size 139x20; Text 'Labeled Bundle'
   TextField "Text field_15" at 145,48 size 84x19; Text 'Pcs'
   TextField "Text field_16" at 228,48 size 87x19; Text '% (From input)'
   TextField "Text field_17" at 7,48 size 139x19; Text 'Output Bundle'
   IOField "I/O field_27" at 253,16 size 66x17; FormatPattern ????????
      ProcessValue <- "Data_String_sDT_Machine id"